   "Carrier_26_SpareSafetyOutput(3_6)" AT %I1665.6 : Bool;   // SPARE SAFETY OUTPUT
   "Carrier_26_SpareSafetyOutput(3_7)" AT %I1665.7 : Bool;   // SPARE SAFETY OUTPUT
   "Carrier_26_Slot4_Input" AT %IW1666 : Word;   // SLOT 4 INPUT WORD
   "Carrier_26_480VPowerOn_MDCB1" AT %I1666.0 : Bool;   // 480 VAC POWER ON MDCB 1
   "Carrier_26_SpareInput(4_1)" AT %I1666.1 : Bool;   // SPARE INPUT
   "Carrier_26_SpareInput(4_2)" AT %I1666.2 : Bool;   // SPARE INPUT
   "Carrier_26_SitopSelectStatus" AT %I1666.3 : Bool;   // SITOP SELECT STATUS
   "Carrier_26_DCsupplyOnPSCB2" AT %I1666.4 : Bool;   // DC SUPPLY ON PSCB 2
   "Carrier_26_SpareInput(4_5)" AT %I1666.5 : Bool;   // SPARE INPUT
   "Carrier_26_SpareInput(4_6)" AT %I1666.6 : Bool;   // SPARE INPUT
   "Carrier_26_SpareInput(4_7)" AT %I1666.7 : Bool;   // SPARE INPUT
   "Carrier_26_PB1_ProdHoldLH" AT %I1667.0 : Bool;   // PB 1 PRODUCTION HOLD LH
   "Carrier_26_PB2_ResetLH" AT %I1667.1 : Bool;   // PB 2 RESET LH
   "Carrier_26_PB3_ProdHoldRH" AT %I1667.2 : Bool;   // PB 3 PRODUCTION HOLD RH
   "Carrier_26_PB4_ResetRH" AT %I1667.3 : Bool;   // PB 4 RESET RH
   "Carrier_26_SpareInput(4_14)" AT %I1667.4 : Bool;   // SPARE INPUT
   "Carrier_26_SpareInput(4_15)" AT %I1667.5 : Bool;   // SPARE INPUT
   "Carrier_26_SpareInput(4_16)" AT %I1667.6 : Bool;   // SPARE INPUT
   "Carrier_26_SpareInput(4_17)" AT %I1667.7 : Bool;   // SPARE INPUT
   "Carrier_26_Slot5_Output" AT %IW1668 : Word;   // SLOT 5 OUTPUT WORD
   "Carrier_26_IRD400_HMI_24VDC_ENABLE" AT %I1668.0 : Bool;   // IRD 400 PANEL HMI 24V DC POWER
   "Carrier_26_FaultLight_LH" AT %I1668.1 : Bool;   // FAULT LIGHT LH
   "Carrier_26_RunLight_LH" AT %I1668.2 : Bool;   // RUN LIGHT LH
   "Carrier_26_FaultLight_RH" AT %I1668.3 : Bool;   // FAULT LIGHT RH
   "Carrier_26_RunLight_RH" AT %I1668.4 : Bool;   // RUN LIGHT RH
   "Carrier_26_SpareOutput(5_5)" AT %I1668.5 : Bool;   // SPARE OUTPUT
   "Carrier_26_SpareOutput(5_6)" AT %I1668.6 : Bool;   // SPARE OUTPUT
   "Carrier_26_SpareOutput(5_7)" AT %I1668.7 : Bool;   // SPARE OUTPUT
   "Carrier_26_ActualSpeed" AT %IW1670 : Word;   // ACTUAL SPEED
   "Carrier_26_CarrierDriveAlarm" AT %IW1672 : Word;   // CARRIER DRIVE ALARM
   "Carrier_26_CarrierDriveWarning" AT %IW1674 : Word;   // CARRIER DRIVE WARNING
   "Carrier_27_Status" AT %IW1700 : Word;   // CARRIER STATUS WORD
   "Carrier_27_Status.0" AT %I1700.0 : Bool;   // HEARTBEAT
   "Carrier_27_Status.1" AT %I1700.1 : Bool;   // MANUAL
   "Carrier_27_Status.2" AT %I1700.2 : Bool;   // IN_AUTO
   "Carrier_27_Status.3" AT %I1700.3 : Bool;   // POSITIONING_COMPLETE
   "Carrier_27_Status.4" AT %I1700.4 : Bool;   // PRODUCTION HOLD
   "Carrier_27_Status.5" AT %I1700.5 : Bool;   // CARRIER MOVING FORWARD
   "Carrier_27_Status.6" AT %I1700.6 : Bool;   // CARRIER MOVING REVERSE
   "Carrier_27_Status.7" AT %I1700.7 : Bool;   // CARRIER FAULT
   "Carrier_27_Status.8" AT %I1701.0 : Bool;   // CRASH DETECT TRIPPED
   "Carrier_27_Status.9" AT %I1701.1 : Bool;
   "Carrier_27_Status.10" AT %I1701.2 : Bool;
   "Carrier_27_Status.11" AT %I1701.3 : Bool;
   "Carrier_27_Status.12" AT %I1701.4 : Bool;
   "Carrier_27_Status.13" AT %I1701.5 : Bool;
   "Carrier_27_Status.14" AT %I1701.6 : Bool;
   "Carrier_27_Status.15" AT %I1701.7 : Bool;
   "Carrier_27_SDCFaultCode" AT %IW1702 : Word;   // SDC FAULT CODE
   "Carrier_27_CarrierPosition" AT %ID1704 : DWord;   // CARRIER POSITION
   "Carrier_27_CarrierNumber" AT %IW1708 : Word;   // CARRIER NUMBER
   "Carrier_27_G120DControlWord" AT %IW1710 : Word;   // G120D_STW1_CONTROL
   "Carrier_27_G120DControlWord.0" AT %I1710.0 : Bool;   // Bit_00_ON
   "Carrier_27_G120DControlWord.1" AT %I1710.1 : Bool;   // Bit_01_AUS2_INH
   "Carrier_27_G120DControlWord.2" AT %I1710.2 : Bool;   // Bit_02_AUS3_STOP
   "Carrier_27_G120DControlWord.3" AT %I1710.3 : Bool;   // Bit_03_EN
   "Carrier_27_G120DControlWord.4" AT %I1710.4 : Bool;   // Bit_04_EN_RAMP
   "Carrier_27_G120DControlWord.5" AT %I1710.5 : Bool;   // Bit_05_START_RAMP
   "Carrier_27_G120DControlWord.6" AT %I1710.6 : Bool;   // Bit_06_SETPOINT
   "Carrier_27_G120DControlWord.7" AT %I1710.7 : Bool;   // Bit_07_RESET
   "Carrier_27_G120DControlWord.8" AT %I1711.0 : Bool;   // Bit_08_JOG_R
   "Carrier_27_G120DControlWord.9" AT %I1711.1 : Bool;   // Bit_09_JOG_L
   "Carrier_27_G120DControlWord.10" AT %I1711.2 : Bool;   // Bit_10_CONTR_PLC
   "Carrier_27_G120DControlWord.11" AT %I1711.3 : Bool;   // Bit_11_REVERSE
   "Carrier_27_G120DControlWord.12" AT %I1711.4 : Bool;   // Bit_12_BRAKE_RELEASE
   "Carrier_27_G120DControlWord.13" AT %I1711.5 : Bool;   // Bit_13_DDS
   "Carrier_27_G120DControlWord.14" AT %I1711.6 : Bool;   // Bit_14_DO0
   "Carrier_27_G120DControlWord.15" AT %I1711.7 : Bool;   // Bit_15_DO1
   "Carrier_27_G120DStatusWord" AT %IW1712 : Word;   // G120D_ZSW1_STATUS
   "Carrier_27_G120DStatusWord.0" AT %I1712.0 : Bool;   // Bit_00_READY_RUN
   "Carrier_27_G120DStatusWord.1" AT %I1712.1 : Bool;   // Bit_01_READY_ON
   "Carrier_27_G120DStatusWord.2" AT %I1712.2 : Bool;   // Bit_02_ENABLE
   "Carrier_27_G120DStatusWord.3" AT %I1712.3 : Bool;   // Bit_03_FAULT
   "Carrier_27_G120DStatusWord.4" AT %I1712.4 : Bool;   // Bit_04_OFF2
   "Carrier_27_G120DStatusWord.5" AT %I1712.5 : Bool;   // Bit_05_OFF3
   "Carrier_27_G120DStatusWord.6" AT %I1712.6 : Bool;   // Bit_06_LOCK_OUT
   "Carrier_27_G120DStatusWord.7" AT %I1712.7 : Bool;   // Bit_07_WARN
   "Carrier_27_G120DStatusWord.8" AT %I1713.0 : Bool;   // Bit_08_NO_DEVIATION
   "Carrier_27_G120DStatusWord.9" AT %I1713.1 : Bool;   // Bit_09_CONTR_PLC
   "Carrier_27_G120DStatusWord.10" AT %I1713.2 : Bool;   // Bit_10_F_MAX
   "Carrier_27_G120DStatusWord.11" AT %I1713.3 : Bool;   // Bit_11_LIMIT_REACHED
   "Carrier_27_G120DStatusWord.12" AT %I1713.4 : Bool;   // Bit_12_BRAKE_OPEN
   "Carrier_27_G120DStatusWord.13" AT %I1713.5 : Bool;   // Bit_13_NO_OVERTEMP
   "Carrier_27_G120DStatusWord.14" AT %I1713.6 : Bool;   // Bit_14_CW_CCW
   "Carrier_27_G120DStatusWord.15" AT %I1713.7 : Bool;   // Bit_15_OVERL
   "Carrier_27_Slot2_Input" AT %IW1714 : Word;   // SLOT 2 INPUT WORD
   "Carrier_27_CrashDetectSW" AT %I1714.0 : Bool;   // CRASH DETECT SW
   "Carrier_27_SpareSafetyInput(2_1)" AT %I1714.1 : Bool;   // SPARE SAFETY INPUT
   "Carrier_27_SpareSafetyInput(2_2)" AT %I1714.2 : Bool;   // SPARE SAFETY INPUT
   "Carrier_27_SpareSafetyInput(2_3)" AT %I1714.3 : Bool;   // SPARE SAFETY INPUT
   "Carrier_27_SpareSafetyInput(2_4)" AT %I1714.4 : Bool;   // SPARE SAFETY INPUT
   "Carrier_27_SpareSafetyInput(2_5)" AT %I1714.5 : Bool;   // SPARE SAFETY INPUT
   "Carrier_27_SpareSafetyInput(2_6)" AT %I1714.6 : Bool;   // SPARE SAFETY INPUT
   "Carrier_27_SpareSafetyInput(2_7)" AT %I1714.7 : Bool;   // SPARE SAFETY INPUT
   "Carrier_27_Slot3_SafetyOutput" AT %IW1715 : Word;   // SLOT 3 SAFETY OUTPUT WORD
   "Carrier_27_Crash_Detect_OK" AT %I1715.0 : Bool;   // CARRIER CRASH DETECT
   "Carrier_27_SpareSafetyOutput(3_1)" AT %I1715.1 : Bool;   // SPARE SAFETY OUTPUT
   "Carrier_27_SpareSafetyOutput(3_2)" AT %I1715.2 : Bool;   // SPARE SAFETY OUTPUT
   "Carrier_27_SpareSafetyOutput(3_3)" AT %I1715.3 : Bool;   // SPARE SAFETY OUTPUT
   "Carrier_27_SpareSafetyOutput(3_4)" AT %I1715.4 : Bool;   // SPARE SAFETY OUTPUT
   "Carrier_27_SpareSafetyOutput(3_5)" AT %I1715.5 : Bool;   // SPARE SAFETY OUTPUT
   "Carrier_27_SpareSafetyOutput(3_6)" AT %I1715.6 : Bool;   // SPARE SAFETY OUTPUT
   "Carrier_27_SpareSafetyOutput(3_7)" AT %I1715.7 : Bool;   // SPARE SAFETY OUTPUT
   "Carrier_27_Slot4_Input" AT %IW1716 : Word;   // SLOT 4 INPUT WORD
   "Carrier_27_480VPowerOn_MDCB1" AT %I1716.0 : Bool;   // 480 VAC POWER ON MDCB 1
   "Carrier_27_SpareInput(4_1)" AT %I1716.1 : Bool;   // SPARE INPUT
   "Carrier_27_SpareInput(4_2)" AT %I1716.2 : Bool;   // SPARE INPUT
   "Carrier_27_SitopSelectStatus" AT %I1716.3 : Bool;   // SITOP SELECT STATUS
   "Carrier_27_DCsupplyOnPSCB2" AT %I1716.4 : Bool;   // DC SUPPLY ON PSCB 2
   "Carrier_27_SpareInput(4_5)" AT %I1716.5 : Bool;   // SPARE INPUT
   "Carrier_27_SpareInput(4_6)" AT %I1716.6 : Bool;   // SPARE INPUT
   "Carrier_27_SpareInput(4_7)" AT %I1716.7 : Bool;   // SPARE INPUT
   "Carrier_27_PB1_ProdHoldLH" AT %I1717.0 : Bool;   // PB 1 PRODUCTION HOLD LH
   "Carrier_27_PB2_ResetLH" AT %I1717.1 : Bool;   // PB 2 RESET LH
   "Carrier_27_PB3_ProdHoldRH" AT %I1717.2 : Bool;   // PB 3 PRODUCTION HOLD RH
   "Carrier_27_PB4_ResetRH" AT %I1717.3 : Bool;   // PB 4 RESET RH
   "Carrier_27_SpareInput(4_14)" AT %I1717.4 : Bool;   // SPARE INPUT
   "Carrier_27_SpareInput(4_15)" AT %I1717.5 : Bool;   // SPARE INPUT
   "Carrier_27_SpareInput(4_16)" AT %I1717.6 : Bool;   // SPARE INPUT
   "Carrier_27_SpareInput(4_17)" AT %I1717.7 : Bool;   // SPARE INPUT
   "Carrier_27_Slot5_Output" AT %IW1718 : Word;   // SLOT 5 OUTPUT WORD
   "Carrier_27_IRD400_HMI_24VDC_ENABLE" AT %I1718.0 : Bool;   // IRD 400 PANEL HMI 24V DC POWER
   "Carrier_27_FaultLight_LH" AT %I1718.1 : Bool;   // FAULT LIGHT LH
   "Carrier_27_RunLight_LH" AT %I1718.2 : Bool;   // RUN LIGHT LH
   "Carrier_27_FaultLight_RH" AT %I1718.3 : Bool;   // FAULT LIGHT RH
   "Carrier_27_RunLight_RH" AT %I1718.4 : Bool;   // RUN LIGHT RH
   "Carrier_27_SpareOutput(5_5)" AT %I1718.5 : Bool;   // SPARE OUTPUT
   "Carrier_27_SpareOutput(5_6)" AT %I1718.6 : Bool;   // SPARE OUTPUT
   "Carrier_27_SpareOutput(5_7)" AT %I1718.7 : Bool;   // SPARE OUTPUT
   "Carrier_27_ActualSpeed" AT %IW1720 : Word;   // ACTUAL SPEED
   "Carrier_27_CarrierDriveAlarm" AT %IW1722 : Word;   // CARRIER DRIVE ALARM
   "Carrier_27_CarrierDriveWarning" AT %IW1724 : Word;   // CARRIER DRIVE WARNING
   "Carrier_28_Status" AT %IW1750 : Word;   // CARRIER STATUS WORD
   "Carrier_28_Status.0" AT %I1750.0 : Bool;   // HEARTBEAT
   "Carrier_28_Status.1" AT %I1750.1 : Bool;   // MANUAL
   "Carrier_28_Status.2" AT %I1750.2 : Bool;   // IN_AUTO
   "Carrier_28_Status.3" AT %I1750.3 : Bool;   // POSITIONING_COMPLETE
   "Carrier_28_Status.4" AT %I1750.4 : Bool;   // PRODUCTION HOLD
   "Carrier_28_Status.5" AT %I1750.5 : Bool;   // CARRIER MOVING FORWARD
   "Carrier_28_Status.6" AT %I1750.6 : Bool;   // CARRIER MOVING REVERSE
   "Carrier_28_Status.7" AT %I1750.7 : Bool;   // CARRIER FAULT
   "Carrier_28_Status.8" AT %I1751.0 : Bool;   // CRASH DETECT TRIPPED
   "Carrier_28_Status.9" AT %I1751.1 : Bool;
   "Carrier_28_Status.10" AT %I1751.2 : Bool;
   "Carrier_28_Status.11" AT %I1751.3 : Bool;
   "Carrier_28_Status.12" AT %I1751.4 : Bool;
   "Carrier_28_Status.13" AT %I1751.5 : Bool;
   "Carrier_28_Status.14" AT %I1751.6 : Bool;
   "Carrier_28_Status.15" AT %I1751.7 : Bool;
   "Carrier_28_SDCFaultCode" AT %IW1752 : Word;   // SDC FAULT CODE
   "Carrier_28_CarrierPosition" AT %ID1754 : DWord;   // CARRIER POSITION
   "Carrier_28_CarrierNumber" AT %IW1758 : Word;   // CARRIER NUMBER
   "Carrier_28_G120DControlWord" AT %IW1760 : Word;   // G120D_STW1_CONTROL
   "Carrier_28_G120DControlWord.0" AT %I1760.0 : Bool;   // Bit_00_ON
   "Carrier_28_G120DControlWord.1" AT %I1760.1 : Bool;   // Bit_01_AUS2_INH
   "Carrier_28_G120DControlWord.2" AT %I1760.2 : Bool;   // Bit_02_AUS3_STOP
   "Carrier_28_G120DControlWord.3" AT %I1760.3 : Bool;   // Bit_03_EN
   "Carrier_28_G120DControlWord.4" AT %I1760.4 : Bool;   // Bit_04_EN_RAMP
   "Carrier_28_G120DControlWord.5" AT %I1760.5 : Bool;   // Bit_05_START_RAMP
   "Carrier_28_G120DControlWord.6" AT %I1760.6 : Bool;   // Bit_06_SETPOINT
   "Carrier_28_G120DControlWord.7" AT %I1760.7 : Bool;   // Bit_07_RESET
   "Carrier_28_G120DControlWord.8" AT %I1761.0 : Bool;   // Bit_08_JOG_R
   "Carrier_28_G120DControlWord.9" AT %I1761.1 : Bool;   // Bit_09_JOG_L
   "Carrier_28_G120DControlWord.10" AT %I1761.2 : Bool;   // Bit_10_CONTR_PLC
   "Carrier_28_G120DControlWord.11" AT %I1761.3 : Bool;   // Bit_11_REVERSE
   "Carrier_28_G120DControlWord.12" AT %I1761.4 : Bool;   // Bit_12_BRAKE_RELEASE
   "Carrier_28_G120DControlWord.13" AT %I1761.5 : Bool;   // Bit_13_DDS
   "Carrier_28_G120DControlWord.14" AT %I1761.6 : Bool;   // Bit_14_DO0
   "Carrier_28_G120DControlWord.15" AT %I1761.7 : Bool;   // Bit_15_DO1
   "Carrier_28_G120DStatusWord" AT %IW1762 : Word;   // G120D_ZSW1_STATUS
   "Carrier_28_G120DStatusWord.0" AT %I1762.0 : Bool;   // Bit_00_READY_RUN
   "Carrier_28_G120DStatusWord.1" AT %I1762.1 : Bool;   // Bit_01_READY_ON
   "Carrier_28_G120DStatusWord.2" AT %I1762.2 : Bool;   // Bit_02_ENABLE
   "Carrier_28_G120DStatusWord.3" AT %I1762.3 : Bool;   // Bit_03_FAULT
   "Carrier_28_G120DStatusWord.4" AT %I1762.4 : Bool;   // Bit_04_OFF2
   "Carrier_28_G120DStatusWord.5" AT %I1762.5 : Bool;   // Bit_05_OFF3
   "Carrier_28_G120DStatusWord.6" AT %I1762.6 : Bool;   // Bit_06_LOCK_OUT
   "Carrier_28_G120DStatusWord.7" AT %I1762.7 : Bool;   // Bit_07_WARN
   "Carrier_28_G120DStatusWord.8" AT %I1763.0 : Bool;   // Bit_08_NO_DEVIATION
   "Carrier_28_G120DStatusWord.9" AT %I1763.1 : Bool;   // Bit_09_CONTR_PLC
   "Carrier_28_G120DStatusWord.10" AT %I1763.2 : Bool;   // Bit_10_F_MAX
   "Carrier_28_G120DStatusWord.11" AT %I1763.3 : Bool;   // Bit_11_LIMIT_REACHED
   "Carrier_28_G120DStatusWord.12" AT %I1763.4 : Bool;   // Bit_12_BRAKE_OPEN
   "Carrier_28_G120DStatusWord.13" AT %I1763.5 : Bool;   // Bit_13_NO_OVERTEMP
   "Carrier_28_G120DStatusWord.14" AT %I1763.6 : Bool;   // Bit_14_CW_CCW
   "Carrier_28_G120DStatusWord.15" AT %I1763.7 : Bool;   // Bit_15_OVERL
   "Carrier_28_Slot2_Input" AT %IW1764 : Word;   // SLOT 2 INPUT WORD
   "Carrier_28_CrashDetectSW" AT %I1764.0 : Bool;   // CRASH DETECT SW
   "Carrier_28_SpareSafetyInput(2_1)" AT %I1764.1 : Bool;   // SPARE SAFETY INPUT
   "Carrier_28_SpareSafetyInput(2_2)" AT %I1764.2 : Bool;   // SPARE SAFETY INPUT
   "Carrier_28_SpareSafetyInput(2_3)" AT %I1764.3 : Bool;   // SPARE SAFETY INPUT
   "Carrier_28_SpareSafetyInput(2_4)" AT %I1764.4 : Bool;   // SPARE SAFETY INPUT
   "Carrier_28_SpareSafetyInput(2_5)" AT %I1764.5 : Bool;   // SPARE SAFETY INPUT
   "Carrier_28_SpareSafetyInput(2_6)" AT %I1764.6 : Bool;   // SPARE SAFETY INPUT
   "Carrier_28_SpareSafetyInput(2_7)" AT %I1764.7 : Bool;   // SPARE SAFETY INPUT
   "Carrier_28_Slot3_SafetyOutput" AT %IW1675 : Word;   // SLOT 3 SAFETY OUTPUT WORD
   "Carrier_28_Crash_Detect_OK" AT %I1675.0 : Bool;   // CARRIER CRASH DETECT
   "Carrier_28_SpareSafetyOutput(3_1)" AT %I1675.1 : Bool;   // SPARE SAFETY OUTPUT
   "Carrier_28_SpareSafetyOutput(3_2)" AT %I1675.2 : Bool;   // SPARE SAFETY OUTPUT
   "Carrier_28_SpareSafetyOutput(3_3)" AT %I1675.3 : Bool;   // SPARE SAFETY OUTPUT
   "Carrier_28_SpareSafetyOutput(3_4)" AT %I1675.4 : Bool;   // SPARE SAFETY OUTPUT
   "Carrier_28_SpareSafetyOutput(3_5)" AT %I1675.5 : Bool;   // SPARE SAFETY OUTPUT
   "Carrier_28_SpareSafetyOutput(3_6)" AT %I1675.6 : Bool;   // SPARE SAFETY OUTPUT
   "Carrier_28_SpareSafetyOutput(3_7)" AT %I1675.7 : Bool;   // SPARE SAFETY OUTPUT
   "Carrier_28_Slot4_Input" AT %IW1766 : Word;   // SLOT 4 INPUT WORD
   "Carrier_28_480VPowerOn_MDCB1" AT %I1766.0 : Bool;   // 480 VAC POWER ON MDCB 1
   "Carrier_28_SpareInput(4_1)" AT %I1766.1 : Bool;   // SPARE INPUT
   "Carrier_28_SpareInput(4_2)" AT %I1766.2 : Bool;   // SPARE INPUT
   "Carrier_28_SitopSelectStatus" AT %I1766.3 : Bool;   // SITOP SELECT STATUS
   "Carrier_28_DCsupplyOnPSCB2" AT %I1766.4 : Bool;   // DC SUPPLY ON PSCB 2
   "Carrier_28_SpareInput(4_5)" AT %I1766.5 : Bool;   // SPARE INPUT
   "Carrier_28_SpareInput(4_6)" AT %I1766.6 : Bool;   // SPARE INPUT
   "Carrier_28_SpareInput(4_7)" AT %I1766.7 : Bool;   // SPARE INPUT
   "Carrier_28_PB1_ProdHoldLH" AT %I1767.0 : Bool;   // PB 1 PRODUCTION HOLD LH
   "Carrier_28_PB2_ResetLH" AT %I1767.1 : Bool;   // PB 2 RESET LH
   "Carrier_28_PB3_ProdHoldRH" AT %I1767.2 : Bool;   // PB 3 PRODUCTION HOLD RH
   "Carrier_28_PB4_ResetRH" AT %I1767.3 : Bool;   // PB 4 RESET RH
   "Carrier_28_SpareInput(4_14)" AT %I1767.4 : Bool;   // SPARE INPUT
   "Carrier_28_SpareInput(4_15)" AT %I1767.5 : Bool;   // SPARE INPUT
   "Carrier_28_SpareInput(4_16)" AT %I1767.6 : Bool;   // SPARE INPUT
   "Carrier_28_SpareInput(4_17)" AT %I1767.7 : Bool;   // SPARE INPUT
   "Carrier_28_Slot5_Output" AT %IW1768 : Word;   // SLOT 5 OUTPUT WORD
   "Carrier_28_IRD400_HMI_24VDC_ENABLE" AT %I1768.0 : Bool;   // IRD 400 PANEL HMI 24V DC POWER
   "Carrier_28_FaultLight_LH" AT %I1768.1 : Bool;   // FAULT LIGHT LH
   "Carrier_28_RunLight_LH" AT %I1768.2 : Bool;   // RUN LIGHT LH
   "Carrier_28_FaultLight_RH" AT %I1768.3 : Bool;   // FAULT LIGHT RH
   "Carrier_28_RunLight_RH" AT %I1768.4 : Bool;   // RUN LIGHT RH
   "Carrier_28_SpareOutput(5_5)" AT %I1768.5 : Bool;   // SPARE OUTPUT
   "Carrier_28_SpareOutput(5_6)" AT %I1768.6 : Bool;   // SPARE OUTPUT
   "Carrier_28_SpareOutput(5_7)" AT %I1768.7 : Bool;   // SPARE OUTPUT
   "Carrier_28_ActualSpeed" AT %IW1770 : Word;   // ACTUAL SPEED
   "Carrier_28_CarrierDriveAlarm" AT %IW1772 : Word;   // CARRIER DRIVE ALARM
   "Carrier_28_CarrierDriveWarning" AT %IW1774 : Word;   // CARRIER DRIVE WARNING
   "Carrier_29_Status" AT %IW1800 : Word;   // CARRIER STATUS WORD
   "Carrier_29_Status.0" AT %I1800.0 : Bool;   // HEARTBEAT
   "Carrier_29_Status.1" AT %I1800.1 : Bool;   // MANUAL
   "Carrier_29_Status.2" AT %I1800.2 : Bool;   // IN_AUTO
   "Carrier_29_Status.3" AT %I1800.3 : Bool;   // POSITIONING_COMPLETE
   "Carrier_29_Status.4" AT %I1800.4 : Bool;   // PRODUCTION HOLD
   "Carrier_29_Status.5" AT %I1800.5 : Bool;   // CARRIER MOVING FORWARD
   "Carrier_29_Status.6" AT %I1800.6 : Bool;   // CARRIER MOVING REVERSE
   "Carrier_29_Status.7" AT %I1800.7 : Bool;   // CARRIER FAULT
   "Carrier_29_Status.8" AT %I1801.0 : Bool;   // CRASH DETECT TRIPPED
   "Carrier_29_Status.9" AT %I1801.1 : Bool;
   "Carrier_29_Status.10" AT %I1801.2 : Bool;
   "Carrier_29_Status.11" AT %I1801.3 : Bool;
   "Carrier_29_Status.12" AT %I1801.4 : Bool;
   "Carrier_29_Status.13" AT %I1801.5 : Bool;
   "Carrier_29_Status.14" AT %I1801.6 : Bool;
   "Carrier_29_Status.15" AT %I1801.7 : Bool;
   "Carrier_29_SDCFaultCode" AT %IW1802 : Word;   // SDC FAULT CODE
   "Carrier_29_CarrierPosition" AT %ID1804 : DWord;   // CARRIER POSITION
   "Carrier_29_CarrierNumber" AT %IW1808 : Word;   // CARRIER NUMBER
   "Carrier_29_G120DControlWord" AT %IW1810 : Word;   // G120D_STW1_CONTROL
   "Carrier_29_G120DControlWord.0" AT %I1810.0 : Bool;   // Bit_00_ON
   "Carrier_29_G120DControlWord.1" AT %I1810.1 : Bool;   // Bit_01_AUS2_INH
   "Carrier_29_G120DControlWord.2" AT %I1810.2 : Bool;   // Bit_02_AUS3_STOP
   "Carrier_29_G120DControlWord.3" AT %I1810.3 : Bool;   // Bit_03_EN
   "Carrier_29_G120DControlWord.4" AT %I1810.4 : Bool;   // Bit_04_EN_RAMP
   "Carrier_29_G120DControlWord.5" AT %I1810.5 : Bool;   // Bit_05_START_RAMP
   "Carrier_29_G120DControlWord.6" AT %I1810.6 : Bool;   // Bit_06_SETPOINT
   "Carrier_29_G120DControlWord.7" AT %I1810.7 : Bool;   // Bit_07_RESET
   "Carrier_29_G120DControlWord.8" AT %I1811.0 : Bool;   // Bit_08_JOG_R
   "Carrier_29_G120DControlWord.9" AT %I1811.1 : Bool;   // Bit_09_JOG_L
   "Carrier_29_G120DControlWord.10" AT %I1811.2 : Bool;   // Bit_10_CONTR_PLC
   "Carrier_29_G120DControlWord.11" AT %I1811.3 : Bool;   // Bit_11_REVERSE
   "Carrier_29_G120DControlWord.12" AT %I1811.4 : Bool;   // Bit_12_BRAKE_RELEASE
   "Carrier_29_G120DControlWord.13" AT %I1811.5 : Bool;   // Bit_13_DDS
   "Carrier_29_G120DControlWord.14" AT %I1811.6 : Bool;   // Bit_14_DO0
   "Carrier_29_G120DControlWord.15" AT %I1811.7 : Bool;   // Bit_15_DO1
   "Carrier_29_G120DStatusWord" AT %IW1812 : Word;   // G120D_ZSW1_STATUS
   "Carrier_29_G120DStatusWord.0" AT %I1812.0 : Bool;   // Bit_00_READY_RUN
   "Carrier_29_G120DStatusWord.1" AT %I1812.1 : Bool;   // Bit_01_READY_ON
   "Carrier_29_G120DStatusWord.2" AT %I1812.2 : Bool;   // Bit_02_ENABLE
   "Carrier_29_G120DStatusWord.3" AT %I1812.3 : Bool;   // Bit_03_FAULT
   "Carrier_29_G120DStatusWord.4" AT %I1812.4 : Bool;   // Bit_04_OFF2
   "Carrier_29_G120DStatusWord.5" AT %I1812.5 : Bool;   // Bit_05_OFF3
   "Carrier_29_G120DStatusWord.6" AT %I1812.6 : Bool;   // Bit_06_LOCK_OUT
   "Carrier_29_G120DStatusWord.7" AT %I1812.7 : Bool;   // Bit_07_WARN
   "Carrier_29_G120DStatusWord.8" AT %I1813.0 : Bool;   // Bit_08_NO_DEVIATION
   "Carrier_29_G120DStatusWord.9" AT %I1813.1 : Bool;   // Bit_09_CONTR_PLC
   "Carrier_29_G120DStatusWord.10" AT %I1813.2 : Bool;   // Bit_10_F_MAX
   "Carrier_29_G120DStatusWord.11" AT %I1813.3 : Bool;   // Bit_11_LIMIT_REACHED
   "Carrier_29_G120DStatusWord.12" AT %I1813.4 : Bool;   // Bit_12_BRAKE_OPEN
   "Carrier_29_G120DStatusWord.13" AT %I1813.5 : Bool;   // Bit_13_NO_OVERTEMP
   "Carrier_29_G120DStatusWord.14" AT %I1813.6 : Bool;   // Bit_14_CW_CCW
   "Carrier_29_G120DStatusWord.15" AT %I1813.7 : Bool;   // Bit_15_OVERL
   "Carrier_29_Slot2_Input" AT %IW1814 : Word;   // SLOT 2 INPUT WORD
   "Carrier_29_CrashDetectSW" AT %I1814.0 : Bool;   // CRASH DETECT SW
   "Carrier_29_SpareSafetyInput(2_1)" AT %I1814.1 : Bool;   // SPARE SAFETY INPUT
   "Carrier_29_SpareSafetyInput(2_2)" AT %I1814.2 : Bool;   // SPARE SAFETY INPUT
   "Carrier_29_SpareSafetyInput(2_3)" AT %I1814.3 : Bool;   // SPARE SAFETY INPUT
   "Carrier_29_SpareSafetyInput(2_4)" AT %I1814.4 : Bool;   // SPARE SAFETY INPUT
   "Carrier_29_SpareSafetyInput(2_5)" AT %I1814.5 : Bool;   // SPARE SAFETY INPUT
   "Carrier_29_SpareSafetyInput(2_6)" AT %I1814.6 : Bool;   // SPARE SAFETY INPUT
   "Carrier_29_SpareSafetyInput(2_7)" AT %I1814.7 : Bool;   // SPARE SAFETY INPUT
   "Carrier_29_Slot3_SafetyOutput" AT %IW1815 : Word;   // SLOT 3 SAFETY OUTPUT WORD
   "Carrier_29_Crash_Detect_OK" AT %I1815.0 : Bool;   // CARRIER CRASH DETECT
   "Carrier_29_SpareSafetyOutput(3_1)" AT %I1815.1 : Bool;   // SPARE SAFETY OUTPUT
   "Carrier_29_SpareSafetyOutput(3_2)" AT %I1815.2 : Bool;   // SPARE SAFETY OUTPUT
   "Carrier_29_SpareSafetyOutput(3_3)" AT %I1815.3 : Bool;   // SPARE SAFETY OUTPUT
   "Carrier_29_SpareSafetyOutput(3_4)" AT %I1815.4 : Bool;   // SPARE SAFETY OUTPUT
   "Carrier_29_SpareSafetyOutput(3_5)" AT %I1815.5 : Bool;   // SPARE SAFETY OUTPUT
   "Carrier_29_SpareSafetyOutput(3_6)" AT %I1815.6 : Bool;   // SPARE SAFETY OUTPUT
   "Carrier_29_SpareSafetyOutput(3_7)" AT %I1815.7 : Bool;   // SPARE SAFETY OUTPUT
   "Carrier_29_Slot4_Input" AT %IW1816 : Word;   // SLOT 4 INPUT WORD
   "Carrier_29_480VPowerOn_MDCB1" AT %I1816.0 : Bool;   // 480 VAC POWER ON MDCB 1
   "Carrier_29_SpareInput(4_1)" AT %I1816.1 : Bool;   // SPARE INPUT
   "Carrier_29_SpareInput(4_2)" AT %I1816.2 : Bool;   // SPARE INPUT
   "Carrier_29_SitopSelectStatus" AT %I1816.3 : Bool;   // SITOP SELECT STATUS
   "Carrier_29_DCsupplyOnPSCB2" AT %I1816.4 : Bool;   // DC SUPPLY ON PSCB 2
   "Carrier_29_SpareInput(4_5)" AT %I1816.5 : Bool;   // SPARE INPUT
   "Carrier_29_SpareInput(4_6)" AT %I1816.6 : Bool;   // SPARE INPUT
   "Carrier_29_SpareInput(4_7)" AT %I1816.7 : Bool;   // SPARE INPUT
   "Carrier_29_PB1_ProdHoldLH" AT %I1817.0 : Bool;   // PB 1 PRODUCTION HOLD LH
   "Carrier_29_PB2_ResetLH" AT %I1817.1 : Bool;   // PB 2 RESET LH
   "Carrier_29_PB3_ProdHoldRH" AT %I1817.2 : Bool;   // PB 3 PRODUCTION HOLD RH
   "Carrier_29_PB4_ResetRH" AT %I1817.3 : Bool;   // PB 4 RESET RH
   "Carrier_29_SpareInput(4_14)" AT %I1817.4 : Bool;   // SPARE INPUT
   "Carrier_29_SpareInput(4_15)" AT %I1817.5 : Bool;   // SPARE INPUT
   "Carrier_29_SpareInput(4_16)" AT %I1817.6 : Bool;   // SPARE INPUT
   "Carrier_29_SpareInput(4_17)" AT %I1817.7 : Bool;   // SPARE INPUT
   "Carrier_29_Slot5_Output" AT %IW1818 : Word;   // SLOT 5 OUTPUT WORD
   "Carrier_29_IRD400_HMI_24VDC_ENABLE" AT %I1818.0 : Bool;   // IRD 400 PANEL HMI 24V DC POWER
   "Carrier_29_FaultLight_LH" AT %I1818.1 : Bool;   // FAULT LIGHT LH
   "Carrier_29_RunLight_LH" AT %I1818.2 : Bool;   // RUN LIGHT LH
   "Carrier_29_FaultLight_RH" AT %I1818.3 : Bool;   // FAULT LIGHT RH
   "Carrier_29_RunLight_RH" AT %I1818.4 : Bool;   // RUN LIGHT RH
   "Carrier_29_SpareOutput(5_5)" AT %I1818.5 : Bool;   // SPARE OUTPUT
   "Carrier_29_SpareOutput(5_6)" AT %I1818.6 : Bool;   // SPARE OUTPUT
   "Carrier_29_SpareOutput(5_7)" AT %I1818.7 : Bool;   // SPARE OUTPUT
   "Carrier_29_ActualSpeed" AT %IW1820 : Word;   // ACTUAL SPEED
   "Carrier_29_CarrierDriveAlarm" AT %IW1822 : Word;   // CARRIER DRIVE ALARM
   "Carrier_29_CarrierDriveWarning" AT %IW1824 : Word;   // CARRIER DRIVE WARNING
   "Carrier_30_Status" AT %IW1850 : Word;   // CARRIER STATUS WORD
   "Carrier_30_Status.0" AT %I1850.0 : Bool;   // HEARTBEAT
   "Carrier_30_Status.1" AT %I1850.1 : Bool;   // MANUAL
   "Carrier_30_Status.2" AT %I1850.2 : Bool;   // IN_AUTO
   "Carrier_30_Status.3" AT %I1850.3 : Bool;   // POSITIONING_COMPLETE
   "Carrier_30_Status.4" AT %I1850.4 : Bool;   // PRODUCTION HOLD
   "Carrier_30_Status.5" AT %I1850.5 : Bool;   // CARRIER MOVING FORWARD
   "Carrier_30_Status.6" AT %I1850.6 : Bool;   // CARRIER MOVING REVERSE
   "Carrier_30_Status.7" AT %I1850.7 : Bool;   // CARRIER FAULT
   "Carrier_30_Status.8" AT %I1851.0 : Bool;   // CRASH DETECT TRIPPED
   "Carrier_30_Status.9" AT %I1851.1 : Bool;
   "Carrier_30_Status.10" AT %I1851.2 : Bool;
   "Carrier_30_Status.11" AT %I1851.3 : Bool;
   "Carrier_30_Status.12" AT %I1851.4 : Bool;
   "Carrier_30_Status.13" AT %I1851.5 : Bool;
   "Carrier_30_Status.14" AT %I1851.6 : Bool;
   "Carrier_30_Status.15" AT %I1851.7 : Bool;
   "Carrier_30_SDCFaultCode" AT %IW1852 : Word;   // SDC FAULT CODE
   "Carrier_30_CarrierPosition" AT %ID1854 : DWord;   // CARRIER POSITION
   "Carrier_30_CarrierNumber" AT %IW1858 : Word;   // CARRIER NUMBER
   "Carrier_30_G120DControlWord" AT %IW1860 : Word;   // G120D_STW1_CONTROL
   "Carrier_30_G120DControlWord.0" AT %I1860.0 : Bool;   // Bit_00_ON
   "Carrier_30_G120DControlWord.1" AT %I1860.1 : Bool;   // Bit_01_AUS2_INH
   "Carrier_30_G120DControlWord.2" AT %I1860.2 : Bool;   // Bit_02_AUS3_STOP
   "Carrier_30_G120DControlWord.3" AT %I1860.3 : Bool;   // Bit_03_EN
   "Carrier_30_G120DControlWord.4" AT %I1860.4 : Bool;   // Bit_04_EN_RAMP
   "Carrier_30_G120DControlWord.5" AT %I1860.5 : Bool;   // Bit_05_START_RAMP
   "Carrier_30_G120DControlWord.6" AT %I1860.6 : Bool;   // Bit_06_SETPOINT
   "Carrier_30_G120DControlWord.7" AT %I1860.7 : Bool;   // Bit_07_RESET
   "Carrier_30_G120DControlWord.8" AT %I1861.0 : Bool;   // Bit_08_JOG_R
   "Carrier_30_G120DControlWord.9" AT %I1861.1 : Bool;   // Bit_09_JOG_L
   "Carrier_30_G120DControlWord.10" AT %I1861.2 : Bool;   // Bit_10_CONTR_PLC
   "Carrier_30_G120DControlWord.11" AT %I1861.3 : Bool;   // Bit_11_REVERSE
   "Carrier_30_G120DControlWord.12" AT %I1861.4 : Bool;   // Bit_12_BRAKE_RELEASE
   "Carrier_30_G120DControlWord.13" AT %I1861.5 : Bool;   // Bit_13_DDS
   "Carrier_30_G120DControlWord.14" AT %I1861.6 : Bool;   // Bit_14_DO0
   "Carrier_30_G120DControlWord.15" AT %I1861.7 : Bool;   // Bit_15_DO1
   "Carrier_30_G120DStatusWord" AT %IW1862 : Word;   // G120D_ZSW1_STATUS
   "Carrier_30_G120DStatusWord.0" AT %I1862.0 : Bool;   // Bit_00_READY_RUN
   "Carrier_30_G120DStatusWord.1" AT %I1862.1 : Bool;   // Bit_01_READY_ON
   "Carrier_30_G120DStatusWord.2" AT %I1862.2 : Bool;   // Bit_02_ENABLE
   "Carrier_30_G120DStatusWord.3" AT %I1862.3 : Bool;   // Bit_03_FAULT
   "Carrier_30_G120DStatusWord.4" AT %I1862.4 : Bool;   // Bit_04_OFF2
   "Carrier_30_G120DStatusWord.5" AT %I1862.5 : Bool;   // Bit_05_OFF3
   "Carrier_30_G120DStatusWord.6" AT %I1862.6 : Bool;   // Bit_06_LOCK_OUT
   "Carrier_30_G120DStatusWord.7" AT %I1862.7 : Bool;   // Bit_07_WARN
   "Carrier_30_G120DStatusWord.8" AT %I1863.0 : Bool;   // Bit_08_NO_DEVIATION
   "Carrier_30_G120DStatusWord.9" AT %I1863.1 : Bool;   // Bit_09_CONTR_PLC
   "Carrier_30_G120DStatusWord.10" AT %I1863.2 : Bool;   // Bit_10_F_MAX
   "Carrier_30_G120DStatusWord.11" AT %I1863.3 : Bool;   // Bit_11_LIMIT_REACHED
   "Carrier_30_G120DStatusWord.12" AT %I1863.4 : Bool;   // Bit_12_BRAKE_OPEN
   "Carrier_30_G120DStatusWord.13" AT %I1863.5 : Bool;   // Bit_13_NO_OVERTEMP
   "Carrier_30_G120DStatusWord.14" AT %I1863.6 : Bool;   // Bit_14_CW_CCW
   "Carrier_30_G120DStatusWord.15" AT %I1863.7 : Bool;   // Bit_15_OVERL
   "Carrier_30_Slot2_Input" AT %IW1864 : Word;   // SLOT 2 INPUT WORD
   "Carrier_30_CrashDetectSW" AT %I1864.0 : Bool;   // CRASH DETECT SW
   "Carrier_30_SpareSafetyInput(2_1)" AT %I1864.1 : Bool;   // SPARE SAFETY INPUT
   "Carrier_30_SpareSafetyInput(2_2)" AT %I1864.2 : Bool;   // SPARE SAFETY INPUT
   "Carrier_30_SpareSafetyInput(2_3)" AT %I1864.3 : Bool;   // SPARE SAFETY INPUT
   "Carrier_30_SpareSafetyInput(2_4)" AT %I1864.4 : Bool;   // SPARE SAFETY INPUT
   "Carrier_30_SpareSafetyInput(2_5)" AT %I1864.5 : Bool;   // SPARE SAFETY INPUT
   "Carrier_30_SpareSafetyInput(2_6)" AT %I1864.6 : Bool;   // SPARE SAFETY INPUT
   "Carrier_30_SpareSafetyInput(2_7)" AT %I1864.7 : Bool;   // SPARE SAFETY INPUT
   "Carrier_30_Slot3_SafetyOutput" AT %IW1685 : Word;   // SLOT 3 SAFETY OUTPUT WORD
   "Carrier_30_Crash_Detect_OK" AT %I1685.0 : Bool;   // CARRIER CRASH DETECT
   "Carrier_30_SpareSafetyOutput(3_1)" AT %I1685.1 : Bool;   // SPARE SAFETY OUTPUT
   "Carrier_30_SpareSafetyOutput(3_2)" AT %I1685.2 : Bool;   // SPARE SAFETY OUTPUT
   "Carrier_30_SpareSafetyOutput(3_3)" AT %I1685.3 : Bool;   // SPARE SAFETY OUTPUT
   "Carrier_30_SpareSafetyOutput(3_4)" AT %I1685.4 : Bool;   // SPARE SAFETY OUTPUT
   "Carrier_30_SpareSafetyOutput(3_5)" AT %I1685.5 : Bool;   // SPARE SAFETY OUTPUT
   "Carrier_30_SpareSafetyOutput(3_6)" AT %I1685.6 : Bool;   // SPARE SAFETY OUTPUT
   "Carrier_30_SpareSafetyOutput(3_7)" AT %I1685.7 : Bool;   // SPARE SAFETY OUTPUT
   "Carrier_30_Slot4_Input" AT %IW1866 : Word;   // SLOT 4 INPUT WORD
   "Carrier_30_480VPowerOn_MDCB1" AT %I1866.0 : Bool;   // 480 VAC POWER ON MDCB 1
   "Carrier_30_SpareInput(4_1)" AT %I1866.1 : Bool;   // SPARE INPUT
   "Carrier_30_SpareInput(4_2)" AT %I1866.2 : Bool;   // SPARE INPUT
   "Carrier_30_SitopSelectStatus" AT %I1866.3 : Bool;   // SITOP SELECT STATUS
   "Carrier_30_DCsupplyOnPSCB2" AT %I1866.4 : Bool;   // DC SUPPLY ON PSCB 2
   "Carrier_30_SpareInput(4_5)" AT %I1866.5 : Bool;   // SPARE INPUT
   "Carrier_30_SpareInput(4_6)" AT %I1866.6 : Bool;   // SPARE INPUT
   "Carrier_30_SpareInput(4_7)" AT %I1866.7 : Bool;   // SPARE INPUT
   "Carrier_30_PB1_ProdHoldLH" AT %I1867.0 : Bool;   // PB 1 PRODUCTION HOLD LH
   "Carrier_30_PB2_ResetLH" AT %I1867.1 : Bool;   // PB 2 RESET LH
   "Carrier_30_PB3_ProdHoldRH" AT %I1867.2 : Bool;   // PB 3 PRODUCTION HOLD RH
   "Carrier_30_PB4_ResetRH" AT %I1867.3 : Bool;   // PB 4 RESET RH
   "Carrier_30_SpareInput(4_14)" AT %I1867.4 : Bool;   // SPARE INPUT
   "Carrier_30_SpareInput(4_15)" AT %I1867.5 : Bool;   // SPARE INPUT
   "Carrier_30_SpareInput(4_16)" AT %I1867.6 : Bool;   // SPARE INPUT
   "Carrier_30_SpareInput(4_17)" AT %I1867.7 : Bool;   // SPARE INPUT
   "Carrier_30_Slot5_Output" AT %IW1868 : Word;   // SLOT 5 OUTPUT WORD
   "Carrier_30_IRD400_HMI_24VDC_ENABLE" AT %I1868.0 : Bool;   // IRD 400 PANEL HMI 24V DC POWER
   "Carrier_30_FaultLight_LH" AT %I1868.1 : Bool;   // FAULT LIGHT LH
   "Carrier_30_RunLight_LH" AT %I1868.2 : Bool;   // RUN LIGHT LH
   "Carrier_30_FaultLight_RH" AT %I1868.3 : Bool;   // FAULT LIGHT RH
   "Carrier_30_RunLight_RH" AT %I1868.4 : Bool;   // RUN LIGHT RH
   "Carrier_30_SpareOutput(5_5)" AT %I1868.5 : Bool;   // SPARE OUTPUT
   "Carrier_30_SpareOutput(5_6)" AT %I1868.6 : Bool;   // SPARE OUTPUT
   "Carrier_30_SpareOutput(5_7)" AT %I1868.7 : Bool;   // SPARE OUTPUT
   "Carrier_30_ActualSpeed" AT %IW1870 : Word;   // ACTUAL SPEED
   "Carrier_30_CarrierDriveAlarm" AT %IW1872 : Word;   // CARRIER DRIVE ALARM
   "Carrier_30_CarrierDriveWarning" AT %IW1874 : Word;   // CARRIER DRIVE WARNING
   "Carrier_31_Status" AT %IW1900 : Word;   // CARRIER STATUS WORD
   "Carrier_31_Status.0" AT %I1900.0 : Bool;   // HEARTBEAT
   "Carrier_31_Status.1" AT %I1900.1 : Bool;   // MANUAL
   "Carrier_31_Status.2" AT %I1900.2 : Bool;   // IN_AUTO
   "Carrier_31_Status.3" AT %I1900.3 : Bool;   // POSITIONING_COMPLETE
   "Carrier_31_Status.4" AT %I1900.4 : Bool;   // PRODUCTION HOLD
   "Carrier_31_Status.5" AT %I1900.5 : Bool;   // CARRIER MOVING FORWARD
   "Carrier_31_Status.6" AT %I1900.6 : Bool;   // CARRIER MOVING REVERSE
   "Carrier_31_Status.7" AT %I1900.7 : Bool;   // CARRIER FAULT
   "Carrier_31_Status.8" AT %I1901.0 : Bool;   // CRASH DETECT TRIPPED
   "Carrier_31_Status.9" AT %I1901.1 : Bool;
   "Carrier_31_Status.10" AT %I1901.2 : Bool;
   "Carrier_31_Status.11" AT %I1901.3 : Bool;
   "Carrier_31_Status.12" AT %I1901.4 : Bool;
   "Carrier_31_Status.13" AT %I1901.5 : Bool;
   "Carrier_31_Status.14" AT %I1901.6 : Bool;
   "Carrier_31_Status.15" AT %I1901.7 : Bool;
   "Carrier_31_SDCFaultCode" AT %IW1902 : Word;   // SDC FAULT CODE
   "Carrier_31_CarrierPosition" AT %ID1904 : DWord;   // CARRIER POSITION
   "Carrier_31_CarrierNumber" AT %IW1908 : Word;   // CARRIER NUMBER
   "Carrier_31_G120DControlWord" AT %IW1910 : Word;   // G120D_STW1_CONTROL
   "Carrier_31_G120DControlWord.0" AT %I1910.0 : Bool;   // Bit_00_ON
   "Carrier_31_G120DControlWord.1" AT %I1910.1 : Bool;   // Bit_01_AUS2_INH
   "Carrier_31_G120DControlWord.2" AT %I1910.2 : Bool;   // Bit_02_AUS3_STOP
   "Carrier_31_G120DControlWord.3" AT %I1910.3 : Bool;   // Bit_03_EN
   "Carrier_31_G120DControlWord.4" AT %I1910.4 : Bool;   // Bit_04_EN_RAMP
   "Carrier_31_G120DControlWord.5" AT %I1910.5 : Bool;   // Bit_05_START_RAMP
   "Carrier_31_G120DControlWord.6" AT %I1910.6 : Bool;   // Bit_06_SETPOINT
   "Carrier_31_G120DControlWord.7" AT %I1910.7 : Bool;   // Bit_07_RESET